text list "Banner_ManIntMsg1": 0 '**Local Message Display**'; 1 '~Spare MB1[0].1'; 2 '~Spare MB1[0].2'; 3 '~Spare MB1[0].3'; 4 '~Spare MB1[0].4'; 5 '~Spare MB1[0].5'; 6 '~Spare MB1[0].6'; 7 '~Spare MB1[0].7'; 8 '~Spare MB1[0].8'; 9 '~Spare MB1[0].9'; 10 '~Spare MB1[0].10'; 11 '~Spare MB1[0].11'; 12 '~Spare MB1[0].12'; 13 '~Spare MB1[0].13'; 14 '~Spare MB1[0].14'; 15 '~Spare MB1[0].15'; 16 '~Spare MB1[0].16'; 17 '~Spare MB1[0].17'; 18 '~Spare MB1[0].18'; 19 '~Spare MB1[0].19'; 20 '~Spare MB1[0].20'; 21 '~Spare MB1[0].21'; 22 '~Spare MB1[0].22'; 23 '~Spare MB1[0].23'; 24 '~Spare MB1[0].24'; 25 '~Spare MB1[0].25'; 26 '~Spare MB1[0].26'; 27 '~Spare MB1[0].27'; 28 '~Spare MB1[0].28'; 29 '~Spare MB1[0].29'; 30 '~Spare MB1[0].30'; 31 '~Spare MB1[0].31'; 32 '~PDPES1 - PDP EtherNet Switch Connection Inhibited MB1[1].0'; 33 '~Spare MB1[1].1'; 34 '~Spare MB1[1].2'; 35 '~MPES1 - Main Panel EtherNet Switch Connection Inhibited MB1[1].3'; 36 '~Spare MB1[1].4'; 37 '~Spare MB1[1].5'; 38 '~MPES2 - Main Panel EtherNet Switch Connection Inhibited MB1[1].6'; 39 '~Spare MB1[1].7'; 40 '~Spare MB1[1].8'; 41 '~MPES3 - Main Panel EtherNet Switch Connection Inhibited MB1[1].9'; 42 '~Spare MB1[1].10'; 43 '~Spare MB1[1].11'; 44 '~S001_004SS1B1 - Service Stand Module Connection Inhibited MB1[1].12'; 45 '~Spare MB1[1].13'; 46 '~Spare MB1[1].14'; 47 '~Spare MB1[1].15'; 48 '~Spare MB1[1].16'; 49 '~MPES1 - Main Panel Control Power Disconnect Not On MB1[1].17'; 50 '~PDP 1 - Panel Output Disconnect Safety Switch Not On MB1[1].18'; 51 '~PDP 2 - Panel Output Disconnect Safety Switch Not On MB1[1].19'; 52 '~PDP 3 - Panel Output Disconnect Safety Switch Not On MB1[1].20'; 53 '~Spare MB1[1].21'; 54 '~Spare MB1[1].22'; 55 '~Spare MB1[1].23'; 56 '~Spare MB1[1].24'; 57 '~Spare MB1[1].25'; 58 '~Spare MB1[1].26'; 59 '~Spare MB1[1].27'; 60 '~Spare MB1[1].28'; 61 '~Spare MB1[1].29'; 62 '~Spare MB1[1].30'; 63 '~Laser Booth-Safe I/O Enclosure Disconnect Safety Switch Not On MB1[1].31'; 64 '~ES1ES1 - ES1 EtherNet Switch Connection Inhibited MB1[2].0'; 65 '~Spare MB1[2].1'; 66 '~Spare MB1[2].2'; 67 '~Spare MB1[2].3'; 68 '~Spare MB1[2].4'; 69 '~Spare MB1[2].5'; 70 '~Spare MB1[2].6'; 71 '~Spare MB1[2].7'; 72 '~Spare MB1[2].8'; 73 '~ES1Sfty - Motion Control Enable Relay #1 MECR1 Still On MB1[2].9'; 74 '~ES1Sfty - Motion Control Enable Relay #1 MECR1 Not On MB1[2].10'; 75 '~ES1Sfty - Motion Control Enable Relay #2 MECR2 Still On MB1[2].11'; 76 '~ES1Sfty - Motion Control Enable Relay #2 MECR2 Not On MB1[2].12'; 77 '~ES1Sfty - EtherNet Switch Sfty Relays RESSR1 RESSR2 Not On MB1[2].13'; 78 '~ES1Sfty - EtherNet Switch Sfty Relays RESSR1 RESSR2 Still On MB1[2].14'; 79 '~Spare MB1[2].15'; 80 '~Spare MB1[2].16'; 81 '~Spare MB1[2].17'; 82 '~Spare MB1[2].18'; 83 '~Spare MB1[2].19'; 84 '~ES1 S001 Safety Gate #1 Open MB1[2].20'; 85 '~ES1 S001 Safety Gate #2 Open MB1[2].21'; 86 '~Spare MB1[2].22'; 87 '~Spare MB1[2].23'; 88 '~Spare MB1[2].24'; 89 '~Spare MB1[2].25'; 90 '~Spare MB1[2].26'; 91 '~Spare MB1[2].27'; 92 '~ES1 S001 Safety Gate #3 Open MB1[2].28'; 93 '~Spare MB1[2].29'; 94 '~Spare MB1[2].30'; 95 '~Spare MB1[2].31'; 96 '~ES2ES1 - ES2 EtherNet Switch Connection Inhibited MB1[3].0'; 97 '~Spare MB1[3].1'; 98 '~Spare MB1[3].2'; 99 '~Spare MB1[3].3'; 100 '~Spare MB1[3].4'; 101 '~Spare MB1[3].5'; 102 '~Spare MB1[3].6'; 103 '~Spare MB1[3].7'; 104 '~Spare MB1[3].8'; 105 '~ES2Sfty - Motion Control Enable Relay #1 MECR1 Still On MB1[3].9'; 106 '~ES2Sfty - Motion Control Enable Relay #1 MECR1 Not On MB1[3].10'; 107 '~ES2Sfty - Motion Control Enable Relay #2 MECR2 Still On MB1[3].11'; 108 '~ES2Sfty - Motion Control Enable Relay #2 MECR2 Not On MB1[3].12'; 109 '~ES2Sfty - EtherNet Switch Sfty Relays RESSR1 RESSR2 Not On MB1[3].13'; 110 '~ES2Sfty - EtherNet Switch Sfty Relays RESSR1 RESSR2 Still On MB1[3].14'; 111 '~Spare MB1[3].15'; 112 '~Spare MB1[3].16'; 113 '~Spare MB1[3].17'; 114 '~Spare MB1[3].18'; 115 '~Spare MB1[3].19'; 116 '~ES2 S001 Safety Gate #1 Open MB1[3].20'; 117 '~ES2 S001 Safety Gate #2 Open MB1[3].21'; 118 '~Spare MB1[3].22'; 119 '~Spare MB1[3].23'; 120 '~Spare MB1[3].24'; 121 '~Spare MB1[3].25'; 122 '~Spare MB1[3].26'; 123 '~Spare MB1[3].27'; 124 '~Spare MB1[3].28'; 125 '~Spare MB1[3].29'; 126 '~Spare MB1[3].30'; 127 '~Spare MB1[3].31'; 128 '~PV1ES1 - PV1 EtherNet Switch Connection Inhibited MB1[4].0'; 129 '~Spare MB1[4].1'; 130 '~Spare MB1[4].2'; 131 '~Spare MB1[4].3'; 132 '~Spare MB1[4].4'; 133 '~Spare MB1[4].5'; 134 '~Spare MB1[4].6'; 135 '~Spare MB1[4].7'; 136 '~Spare MB1[4].8'; 137 '~Spare MB1[4].9'; 138 '~Spare MB1[4].10'; 139 '~PV1Sfty - EtherNet Switch Sfty Relays RESSR1 RESSR2 Not On MB1[4].11'; 140 '~PV1Sfty - EtherNet Switch Sfty Relays RESSR1 RESSR2 Still On MB1[4].12'; 141 '~Spare MB1[4].13'; 142 '~Spare MB1[4].14'; 143 '~PV1 S001 E-Stop Depressed MB1[4].15'; 144 '~PV1 S001 Safety Gate #1 Open MB1[4].16'; 145 '~PV1 S001 Safety Gate #2 Open MB1[4].17'; 146 '~PV1 S001 Safety Gate #3 Open MB1[4].18'; 147 '~Spare MB1[4].19'; 148 '~Spare MB1[4].20'; 149 '~Spare MB1[4].21'; 150 '~Spare MB1[4].22'; 151 '~Spare MB1[4].23'; 152 '~S001 Both PanelViews Have Manual Selected MB1[4].24'; 153 '~S001 PanelView 1 Manual Selected MB1[4].25'; 154 '~Spare MB1[4].26'; 155 '~Spare MB1[4].27'; 156 '~PV1 S001 Auto Not Selected MB1[4].28'; 157 '~PV1 S001 Not In Auto Or Manual MB1[4].29'; 158 '~Spare MB1[4].30'; 159 '~Spare MB1[4].31'; 160 '~PV2ES1 - PV2 EtherNet Switch Connection Inhibited MB1[5].0'; 161 '~Spare MB1[5].1'; 162 '~Spare MB1[5].2'; 163 '~Spare MB1[5].3'; 164 '~Spare MB1[5].4'; 165 '~Spare MB1[5].5'; 166 '~Spare MB1[5].6'; 167 '~Spare MB1[5].7'; 168 '~Spare MB1[5].8'; 169 '~Spare MB1[5].9'; 170 '~Spare MB1[5].10'; 171 '~PV2Sfty - EtherNet Switch Sfty Relays RESSR1 RESSR2 Not On MB1[5].11'; 172 '~PV2Sfty - EtherNet Switch Sfty Relays RESSR1 RESSR2 Still On MB1[5].12'; 173 '~Spare MB1[5].13'; 174 '~Spare MB1[5].14'; 175 '~PV2 S001 E-Stop Depressed MB1[5].15'; 176 '~PV2 S001 Safety Gate #1 Open MB1[5].16'; 177 '~PV2 S001 Safety Gate #2 Open MB1[5].17'; 178 '~PV2 S001 Safety Gate #3 Open MB1[5].18'; 179 '~Spare MB1[5].19'; 180 '~Spare MB1[5].20'; 181 '~Spare MB1[5].21'; 182 '~Spare MB1[5].22'; 183 '~Spare MB1[5].23'; 184 '~Spare MB1[5].24'; 185 '~S001 PanelView 2 Manual Selected MB1[5].25'; 186 '~Spare MB1[5].26'; 187 '~Spare MB1[5].27'; 188 '~PV2 S001 Auto Not Selected MB1[5].28'; 189 '~PV2 S001 Not In Auto Or Manual MB1[5].29'; 190 '~Spare MB1[5].30'; 191 '~Spare MB1[5].31'; 192 '~S001R01ES1 - S001R01 EtherNet Switch Connection Inhibited MB1[6].0'; 193 '~Spare MB1[6].1'; 194 '~Spare MB1[6].2'; 195 '~Spare MB1[6].3'; 196 '~Spare MB1[6].4'; 197 '~Spare MB1[6].5'; 198 '~Spare MB1[6].6'; 199 '~Spare MB1[6].7'; 200 '~Spare MB1[6].8'; 201 '~Spare MB1[6].9'; 202 '~Spare MB1[6].10'; 203 '~Spare MB1[6].11'; 204 '~Spare MB1[6].12'; 205 '~Spare MB1[6].13'; 206 '~Spare MB1[6].14'; 207 '~Spare MB1[6].15'; 208 '~Spare MB1[6].16'; 209 '~S001R01Sfty - Robot E-Stop Depressed MB1[6].17'; 210 '~S001R01Sfty - Robot Safety Interface Not Enabled MB1[6].18'; 211 '~S001R01Sfty - Robot DCS Has Been Edited MB1[6].19'; 212 '~S001R01CN - Robot Controller Connection Inhibited MB1[6].20'; 213 '~S001R01E#B# - Robot End Effector Module Connection Inhibited MB1[6].21'; 214 '~S001R01E#B# - Robot End Effector Module Connection Inhibited MB1[6].22'; 215 '~S001R01E#B# - Robot End Effector Module Connection Inhibited MB1[6].23'; 216 '~S001R01E#B# - Robot End Effector Module Connection Inhibited MB1[6].24'; 217 '~S001R01E#B# - Robot End Effector Module Connection Inhibited MB1[6].25'; 218 '~S001R01E#B# - Robot End Effector Module Connection Inhibited MB1[6].26'; 219 '~S001R01E#B# - Robot End Effector Module Connection Inhibited MB1[6].27'; 220 '~S001R01E#B# - Robot End Effector Module Connection Inhibited MB1[6].28'; 221 '~S001R01E#B# - Robot End Effector Module Connection Inhibited MB1[6].29'; 222 '~Spare MB1[6].30'; 223 '~Spare MB1[6].31'; 224 '~Spare MB1[7].0'; 225 '~S001R01F#B# - Robot Process I/O Connection Inhibited MB1[7].1'; 226 '~S001R01F#B# - Robot Process I/O Connection Inhibited MB1[7].2'; 227 '~S001R01F#B# - Robot Process I/O Connection Inhibited MB1[7].3'; 228 '~S001R01F#B# - Robot Process I/O Connection Inhibited MB1[7].4'; 229 '~Spare MB1[7].5'; 230 '~Spare MB1[7].6'; 231 '~Spare MB1[7].7'; 232 '~Spare MB1[7].8'; 233 '~Spare MB1[7].9'; 234 '~S001R01CN.I.Safety - Chain Fault MB1[7].10'; 235 '~S001R01CN.I.AirOn - Robot Air Not On MB1[7].11'; 236 '~S001R01CN.I.RbtAuto - Robot Not in Auto MB1[7].12'; 237 '~S001R01CN.M.InTeach - Robot In Teach MB1[7].13'; 238 '~S001R01CN.I.AtMaintPos - Robot At Maintenace MB1[7].14'; 239 '~S001R01CN.I.RunEnblInterruptAck - Robot In Hold MB1[7].15'; 240 '~S001R01CN.M.MaintPosSeld - Robot Maintenance Selected MB1[7].16'; 241 '~Spare MB1[7].17'; 242 '~Spare MB1[7].18'; 243 '~Spare MB1[7].19'; 244 '~S001R01CN.I.ExtAppCommFlt - Robot Application Communication Fault MB1[7].20'; 245 '~S001R01CN.M.AbortPickupSeld - Robot Abort Pickup Selected MB1[7].21'; 246 '~S001R01CN.M.RetFmPounceSeld - Robot Return From Pounce Selected MB1[7].22'; 247 '~S001R01CN.I.StudWld1 Comm Not OK MB1[7].23'; 248 '~S001R01CN.I.StudWld2 Comm Not OK MB1[7].24'; 249 '~S001R01CN.I.WldMode - Robot In No Weld MB1[7].25'; 250 '~S001R01CN.I.PulledTipBypSS - Robot Pulled Tip Bypass Selected MB1[7].26'; 251 '~S001R01CN.I.FlowNoFlowSS - Robot In No Flow MB1[7].27'; 252 '~S001R01CN.I.RvtNoRvtSS - Robot In No Rivet MB1[7].28'; 253 '~S001R01CN.I.WldCtrlCommOk1 - Robot Weld Controller 1 Comm Not OK MB1[7].29'; 254 '~S001R01CN.I.WldModeStud - Robot In No Weld Stud MB1[7].30'; 255 '~S001R01CN.Ix.MigWldNoWld - Robot In No Weld Mig MB1[7].31'; 256 '~S001R01CN.I.StudWld1Rdy - Robot Stud Weld Controller 1 Not Ready MB1[8].0'; 257 '~S001R01CN.I.Rvt1RdyToOperate - Robot Rivet Controller 1 Not Ready MB1[8].1'; 258 '~S001R01CN.Ix.MigRdy - Robot Mig Weld Controller Not Ready MB1[8].2'; 259 '~S001R01CN.Ix.MigWldNoWld - Robot In No Weld MB1[8].3'; 260 '~Spare MB1[8].4'; 261 '~S001R01CN.I.WldCtrlCommOk2 - Robot Weld Controller 2 Comm Not OK MB1[8].5'; 262 '~Spare MB1[8].6'; 263 '~Spare MB1[8].7'; 264 '~S001R01CN.I.StudWld2Rdy - Robot Stud Weld Controller 2 Not Ready MB1[8].8'; 265 '~S001R01CN.I.Rvt2RdyToOperate - Robot Rivet Controller 2 Not Ready MB1[8].9'; 266 '~S001R01CN.Ix.LaserWldOn - Robot Laser In No Cut MB1[8].10'; 267 '~S001R01CN.Ix.GlassNotPres - Robot Laser Glass Not Present MB1[8].11'; 268 '~S001R01CN.Ix.LaserHeadRdy - Robot Laser Head Not Ready MB1[8].12'; 269 '~S001R01CN.Ix.ChillerOn - Robot Laser Chiller Not On MB1[8].13'; 270 '~S001R01CN.Ix.GasOn - Robot Gas Not On MB1[8].14'; 271 '~S001R01 Power Meter Not Ready MB1[8].15'; 272 '~S001R01 No Wire Present Replace Barrel MB1[8].16'; 273 '~S001R01 Wire Feeder Fault Timer MB1[8].17'; 274 '~S001R01CN.Ix.NRFlt - Robot Nut Runner Not Ready MB1[8].18'; 275 '~Spare MB1[8].19'; 276 '~S001R01CN.M.WrongRivetAtNose - Remove Wrong Rivet At Nose MB1[8].20'; 277 '~S001R01CN.M.DisableRbtDrvs - In Rivet Zone But Riveter Not In Auto MB1[8].21'; 278 '~S001R01CN.I.Rvt1SystemInAuto - Rivet Controller 1 Not In Auto MB1[8].22'; 279 '~S001R01CN.I.Rvt2SystemInAuto - Rivet Controller 2 Not In Auto MB1[8].23'; 280 '~S001R01CN.M.RvtC1ReelCtr.DN - Reel Change Required MB1[8].24'; 281 '~S001R01CN.M.RvtC2ReelCtr.DN - Reel Change Required MB1[8].25'; 282 '~S001R01CN.M.AbortSkipRemain - SkipRemaining Aborted, Reset At Rbt Controller Is Required MB1[8].26'; 283 '~Spare MB1[8].27'; 284 '~Spare MB1[8].28'; 285 '~Spare MB1[8].29'; 286 '~Spare MB1[8].30'; 287 '~Spare MB1[8].31'; 288 '~Spare MB1[9].0'; 289 '~Spare MB1[9].1'; 290 '~Spare MB1[9].2'; 291 '~Spare MB1[9].3'; 292 '~Spare MB1[9].4'; 293 '~Spare MB1[9].5'; 294 '~Spare MB1[9].6'; 295 '~Spare MB1[9].7'; 296 '~Spare MB1[9].8'; 297 '~Spare MB1[9].9'; 298 '~Spare MB1[9].10'; 299 '~Spare MB1[9].11'; 300 '~Spare MB1[9].12'; 301 '~Spare MB1[9].13'; 302 '~Spare MB1[9].14'; 303 '~Spare MB1[9].15'; 304 '~Spare MB1[9].16'; 305 '~Spare MB1[9].17'; 306 '~Spare MB1[9].18'; 307 '~Spare MB1[9].19'; 308 '~Spare MB1[9].20'; 309 '~Spare MB1[9].21'; 310 '~Spare MB1[9].22'; 311 '~Spare MB1[9].23'; 312 '~Spare MB1[9].24'; 313 '~Spare MB1[9].25'; 314 '~Spare MB1[9].26'; 315 '~Spare MB1[9].27'; 316 '~Spare MB1[9].28'; 317 '~Spare MB1[9].29'; 318 '~Spare MB1[9].30'; 319 '~Spare MB1[9].31'; 320 '~Spare MB1[10].0'; 321 '~Spare MB1[10].1'; 322 '~Spare MB1[10].2'; 323 '~Spare MB1[10].3'; 324 '~Spare MB1[10].4'; 325 '~Spare MB1[10].5'; 326 '~Spare MB1[10].6'; 327 '~Spare MB1[10].7'; 328 '~Spare MB1[10].8'; 329 '~Spare MB1[10].9'; 330 '~Spare MB1[10].10'; 331 '~Spare MB1[10].11'; 332 '~Spare MB1[10].12'; 333 '~Spare MB1[10].13'; 334 '~Spare MB1[10].14'; 335 '~Spare MB1[10].15'; 336 '~Spare MB1[10].16'; 337 '~Spare MB1[10].17'; 338 '~Spare MB1[10].18'; 339 '~Spare MB1[10].19'; 340 '~Spare MB1[10].20'; 341 '~Spare MB1[10].21'; 342 '~Spare MB1[10].22'; 343 '~Spare MB1[10].23'; 344 '~Spare MB1[10].24'; 345 '~Spare MB1[10].25'; 346 '~Spare MB1[10].26'; 347 '~Spare MB1[10].27'; 348 '~Spare MB1[10].28'; 349 '~Spare MB1[10].29'; 350 '~Spare MB1[10].30'; 351 '~Spare MB1[10].31'; 352 '~Spare MB1[11].0'; 353 '~Spare MB1[11].1'; 354 '~Spare MB1[11].2'; 355 '~Spare MB1[11].3'; 356 '~Spare MB1[11].4'; 357 '~Spare MB1[11].5'; 358 '~Spare MB1[11].6'; 359 '~Spare MB1[11].7'; 360 '~Spare MB1[11].8'; 361 '~Spare MB1[11].9'; 362 '~Spare MB1[11].10'; 363 '~Spare MB1[11].11'; 364 '~Spare MB1[11].12'; 365 '~Spare MB1[11].13'; 366 '~Spare MB1[11].14'; 367 '~Spare MB1[11].15'; 368 '~Spare MB1[11].16'; 369 '~Spare MB1[11].17'; 370 '~Spare MB1[11].18'; 371 '~Spare MB1[11].19'; 372 '~Spare MB1[11].20'; 373 '~Spare MB1[11].21'; 374 '~Spare MB1[11].22'; 375 '~Spare MB1[11].23'; 376 '~Spare MB1[11].24'; 377 '~Spare MB1[11].25'; 378 '~Spare MB1[11].26'; 379 '~Spare MB1[11].27'; 380 '~Spare MB1[11].28'; 381 '~Spare MB1[11].29'; 382 '~Spare MB1[11].30'; 383 '~Spare MB1[11].31'; 384 '~S001R02ES1 - S001R02 EtherNet Switch Connection Inhibited MB1[12].0'; 385 '~Spare MB1[12].1'; 386 '~Spare MB1[12].2'; 387 '~Spare MB1[12].3'; 388 '~Spare MB1[12].4'; 389 '~Spare MB1[12].5'; 390 '~Spare MB1[12].6'; 391 '~Spare MB1[12].7'; 392 '~Spare MB1[12].8'; 393 '~Spare MB1[12].9'; 394 '~Spare MB1[12].10'; 395 '~Spare MB1[12].11'; 396 '~Spare MB1[12].12'; 397 '~Spare MB1[12].13'; 398 '~Spare MB1[12].14'; 399 '~Spare MB1[12].15'; 400 '~Spare MB1[12].16'; 401 '~S001R02Sfty - Robot E-Stop Depressed MB1[12].17'; 402 '~S001R02Sfty - Robot Safety Interface Not Enabled MB1[12].18'; 403 '~S001R02Sfty - Robot DCS Has Been Edited MB1[12].19'; 404 '~S001R02CN - Robot Controller Connection Inhibited MB1[12].20'; 405 '~S001R02E#B# - Robot End Effector Module Connection Inhibited MB1[12].21'; 406 '~S001R02E#B# - Robot End Effector Module Connection Inhibited MB1[12].22'; 407 '~S001R02E#B# - Robot End Effector Module Connection Inhibited MB1[12].23'; 408 '~S001R02E#B# - Robot End Effector Module Connection Inhibited MB1[12].24'; 409 '~S001R02E#B# - Robot End Effector Module Connection Inhibited MB1[12].25'; 410 '~S001R02E#B# - Robot End Effector Module Connection Inhibited MB1[12].26'; 411 '~S001R02E#B# - Robot End Effector Module Connection Inhibited MB1[12].27'; 412 '~S001R02E#B# - Robot End Effector Module Connection Inhibited MB1[12].28'; 413 '~S001R02E#B# - Robot End Effector Module Connection Inhibited MB1[12].29'; 414 '~Spare MB1[12].30'; 415 '~Spare MB1[12].31'; 416 '~Spare MB1[13].0'; 417 '~S001R02F#B# - Robot Process I/O Connection Inhibited MB1[13].1'; 418 '~S001R02F#B# - Robot Process I/O Connection Inhibited MB1[13].2'; 419 '~S001R02F#B# - Robot Process I/O Connection Inhibited MB1[13].3'; 420 '~S001R02F#B# - Robot Process I/O Connection Inhibited MB1[13].4'; 421 '~Spare MB1[13].5'; 422 '~Spare MB1[13].6'; 423 '~Spare MB1[13].7'; 424 '~Spare MB1[13].8'; 425 '~Spare MB1[13].9'; 426 '~S001R02CN.I.Safety - Chain Fault MB1[13].10'; 427 '~S001R02CN.I.AirOn - Robot Air Not On MB1[13].11'; 428 '~S001R02CN.I.RbtAuto - Robot Not in Auto MB1[13].12'; 429 '~S001R02CN.M.InTeach - Robot In Teach MB1[13].13'; 430 '~S001R02CN.I.AtMaintPos - Robot At Maintenace MB1[13].14'; 431 '~S001R02CN.I.RunEnblInterruptAck - Robot In Hold MB1[13].15'; 432 '~S001R02CN.M.MaintPosSeld - Robot Maintenance Selected MB1[13].16'; 433 '~Spare MB1[13].17'; 434 '~Spare MB1[13].18'; 435 '~Spare MB1[13].19'; 436 '~S001R02CN.I.ExtAppCommFlt - Robot Application Communication Fault MB1[13].20'; 437 '~S001R02CN.M.AbortPickupSeld - Robot Abort Pickup Selected MB1[13].21'; 438 '~S001R02CN.M.RetFmPounceSeld - Robot Return From Pounce Selected MB1[13].22'; 439 '~S001R02CN.I.StudWld1 Comm Not OK MB1[13].23'; 440 '~S001R02CN.I.StudWld2 Comm Not OK MB1[13].24'; 441 '~S001R02CN.I.WldMode - Robot In No Weld MB1[13].25'; 442 '~S001R02CN.I.PulledTipBypSS - Robot Pulled Tip Bypass Selected MB1[13].26'; 443 '~S001R02CN.I.FlowNoFlowSS - Robot In No Flow MB1[13].27'; 444 '~S001R02CN.I.RvtNoRvtSS - Robot In No Rivet MB1[13].28'; 445 '~S001R02CN.I.WldCtrlCommOk1 - Robot Weld Controller 1 Comm Not OK MB1[13].29'; 446 '~S001R02CN.I.WldModeStud - Robot In No Weld Stud MB1[13].30'; 447 '~S001R02CN.Ix.MigWldNoWld - Robot In No Weld Mig MB1[13].31'; 448 '~S001R02CN.I.StudWld1Rdy - Robot Stud Weld Controller 1 Not Ready MB1[14].0'; 449 '~S001R02CN.I.Rvt1RdyToOperate - Robot Rivet Controller 1 Not Ready MB1[14].1'; 450 '~S001R02CN.Ix.MigRdy - Robot Mig Weld Controller Not Ready MB1[14].2'; 451 '~S001R02CN.Ix.MigWldNoWld - Robot In No Weld MB1[14].3'; 452 '~Spare MB1[14].4'; 453 '~S001R02CN.I.WldCtrlCommOk2 - Robot Weld Controller 2 Comm Not OK MB1[14].5'; 454 '~Spare MB1[14].6'; 455 '~Spare MB1[14].7'; 456 '~S001R02CN.I.StudWld2Rdy - Robot Stud Weld Controller 2 Not Ready MB1[14].8'; 457 '~S001R02CN.I.Rvt2RdyToOperate - Robot Rivet Controller 2 Not Ready MB1[14].9'; 458 '~S001R02CN.Ix.LaserWldOn - Robot Laser In No Cut MB1[14].10'; 459 '~S001R02CN.Ix.GlassNotPres - Robot Laser Glass Not Present MB1[14].11'; 460 '~S001R02CN.Ix.LaserHeadRdy - Robot Laser Head Not Ready MB1[14].12'; 461 '~S001R02CN.Ix.ChillerOn - Robot Laser Chiller Not On MB1[14].13'; 462 '~S001R02CN.Ix.GasOn - Robot Gas Not On MB1[14].14'; 463 '~S001R02 Power Meter Not Ready MB1[14].15'; 464 '~S001R02 No Wire Present Replace Barrel MB1[14].16'; 465 '~S001R02 Wire Feeder Fault Timer MB1[14].17'; 466 '~S001R02CN.Ix.NRFlt - Robot Nut Runner Not Ready MB1[14].18'; 467 '~Spare MB1[14].19'; 468 '~S001R02CN.M.WrongRivetAtNose - Remove Wrong Rivet At Nose MB1[14].20'; 469 '~S001R02CN.M.DisableRbtDrvs - In Rivet Zone But Riveter Not In Auto MB1[14].21'; 470 '~S001R02CN.I.Rvt1SystemInAuto - Rivet Controller 1 Not In Auto MB1[14].22'; 471 '~S001R02CN.I.Rvt2SystemInAuto - Rivet Controller 2 Not In Auto MB1[14].23'; 472 '~S001R02CN.M.RvtC1ReelCtr.DN - Reel Change Required MB1[14].24'; 473 '~S001R02CN.M.RvtC2ReelCtr.DN - Reel Change Required MB1[14].25'; 474 '~S001R02CN.M.AbortSkipRemain - SkipRemaining Aborted, Reset At Rbt Controller Is Required MB1[14].26'; 475 '~Spare MB1[14].27'; 476 '~Spare MB1[14].28'; 477 '~Spare MB1[14].29'; 478 '~Spare MB1[14].30'; 479 '~Spare MB1[14].31'; 480 '~Spare MB1[15].0'; 481 '~Spare MB1[15].1'; 482 '~Spare MB1[15].2'; 483 '~Spare MB1[15].3'; 484 '~Spare MB1[15].4'; 485 '~Spare MB1[15].5'; 486 '~Spare MB1[15].6'; 487 '~Spare MB1[15].7'; 488 '~Spare MB1[15].8'; 489 '~Spare MB1[15].9'; 490 '~Spare MB1[15].10'; 491 '~Spare MB1[15].11'; 492 '~Spare MB1[15].12'; 493 '~Spare MB1[15].13'; 494 '~Spare MB1[15].14'; 495 '~Spare MB1[15].15'; 496 '~Spare MB1[15].16'; 497 '~Spare MB1[15].17'; 498 '~Spare MB1[15].18'; 499 '~Spare MB1[15].19'; 500 '~Spare MB1[15].20'; 501 '~Spare MB1[15].21'; 502 '~Spare MB1[15].22'; 503 '~Spare MB1[15].23'; 504 '~Spare MB1[15].24'; 505 '~Spare MB1[15].25'; 506 '~Spare MB1[15].26'; 507 '~Spare MB1[15].27'; 508 '~Spare MB1[15].28'; 509 '~Spare MB1[15].29'; 510 '~Spare MB1[15].30'; 511 '~Spare MB1[15].31'; 512 '~Spare MB1[16].0'; 513 '~Spare MB1[16].1'; 514 '~Spare MB1[16].2'; 515 '~Spare MB1[16].3'; 516 '~Spare MB1[16].4'; 517 '~Spare MB1[16].5'; 518 '~Spare MB1[16].6'; 519 '~Spare MB1[16].7'; 520 '~Spare MB1[16].8'; 521 '~Spare MB1[16].9'; 522 '~Spare MB1[16].10'; 523 '~Spare MB1[16].11'; 524 '~Spare MB1[16].12'; 525 '~Spare MB1[16].13'; 526 '~Spare MB1[16].14'; 527 '~Spare MB1[16].15'; 528 '~Spare MB1[16].16'; 529 '~Spare MB1[16].17'; 530 '~Spare MB1[16].18'; 531 '~Spare MB1[16].19'; 532 '~Spare MB1[16].20'; 533 '~Spare MB1[16].21'; 534 '~Spare MB1[16].22'; 535 '~Spare MB1[16].23'; 536 '~Spare MB1[16].24'; 537 '~Spare MB1[16].25'; 538 '~Spare MB1[16].26'; 539 '~Spare MB1[16].27'; 540 '~Spare MB1[16].28'; 541 '~Spare MB1[16].29'; 542 '~Spare MB1[16].30'; 543 '~Spare MB1[16].31'; 544 '~Spare MB1[17].0'; 545 '~Spare MB1[17].1'; 546 '~Spare MB1[17].2'; 547 '~Spare MB1[17].3'; 548 '~Spare MB1[17].4'; 549 '~Spare MB1[17].5'; 550 '~Spare MB1[17].6'; 551 '~Spare MB1[17].7'; 552 '~Spare MB1[17].8'; 553 '~Spare MB1[17].9'; 554 '~Spare MB1[17].10'; 555 '~Spare MB1[17].11'; 556 '~Spare MB1[17].12'; 557 '~Spare MB1[17].13'; 558 '~Spare MB1[17].14'; 559 '~Spare MB1[17].15'; 560 '~Spare MB1[17].16'; 561 '~Spare MB1[17].17'; 562 '~Spare MB1[17].18'; 563 '~Spare MB1[17].19'; 564 '~Spare MB1[17].20'; 565 '~Spare MB1[17].21'; 566 '~Spare MB1[17].22'; 567 '~Spare MB1[17].23'; 568 '~Spare MB1[17].24'; 569 '~Spare MB1[17].25'; 570 '~Spare MB1[17].26'; 571 '~Spare MB1[17].27'; 572 '~Spare MB1[17].28'; 573 '~Spare MB1[17].29'; 574 '~Spare MB1[17].30'; 575 '~Spare MB1[17].31'; 576 '~S001R03ES1 - S001R03 EtherNet Switch Connection Inhibited MB1[18].0'; 577 '~Spare MB1[18].1'; 578 '~Spare MB1[18].2'; 579 '~Spare MB1[18].3'; 580 '~Spare MB1[18].4'; 581 '~Spare MB1[18].5'; 582 '~Spare MB1[18].6'; 583 '~Spare MB1[18].7'; 584 '~Spare MB1[18].8'; 585 '~Spare MB1[18].9'; 586 '~Spare MB1[18].10'; 587 '~Spare MB1[18].11'; 588 '~Spare MB1[18].12'; 589 '~Spare MB1[18].13'; 590 '~Spare MB1[18].14'; 591 '~Spare MB1[18].15'; 592 '~Spare MB1[18].16'; 593 '~S001R03Sfty - Robot E-Stop Depressed MB1[18].17'; 594 '~S001R03Sfty - Robot Safety Interface Not Enabled MB1[18].18'; 595 '~S001R03Sfty - Robot DCS Has Been Edited MB1[18].19'; 596 '~S001R03CN - Robot Controller Connection Inhibited MB1[18].20'; 597 '~S001R03E#B# - Robot End Effector Module Connection Inhibited MB1[18].21'; 598 '~S001R03E#B# - Robot End Effector Module Connection Inhibited MB1[18].22'; 599 '~S001R03E#B# - Robot End Effector Module Connection Inhibited MB1[18].23'; 600 '~S001R03E#B# - Robot End Effector Module Connection Inhibited MB1[18].24'; 601 '~S001R03E#B# - Robot End Effector Module Connection Inhibited MB1[18].25'; 602 '~S001R03E#B# - Robot End Effector Module Connection Inhibited MB1[18].26'; 603 '~S001R03E#B# - Robot End Effector Module Connection Inhibited MB1[18].27'; 604 '~S001R03E#B# - Robot End Effector Module Connection Inhibited MB1[18].28'; 605 '~S001R03E#B# - Robot End Effector Module Connection Inhibited MB1[18].29'; 606 '~Spare MB1[18].30'; 607 '~Spare MB1[18].31'; 608 '~Spare MB1[19].0'; 609 '~S001R03F#B# - Robot Process I/O Connection Inhibited MB1[19].1'; 610 '~S001R03F#B# - Robot Process I/O Connection Inhibited MB1[19].2'; 611 '~S001R03F#B# - Robot Process I/O Connection Inhibited MB1[19].3'; 612 '~S001R03F#B# - Robot Process I/O Connection Inhibited MB1[19].4'; 613 '~Spare MB1[19].5'; 614 '~Spare MB1[19].6'; 615 '~Spare MB1[19].7'; 616 '~Spare MB1[19].8'; 617 '~Spare MB1[19].9'; 618 '~S001R03CN.I.Safety - Chain Fault MB1[19].10'; 619 '~S001R03CN.I.AirOn - Robot Air Not On MB1[19].11'; 620 '~S001R03CN.I.RbtAuto - Robot Not in Auto MB1[19].12'; 621 '~S001R03CN.M.InTeach - Robot In Teach MB1[19].13'; 622 '~S001R03CN.I.AtMaintPos - Robot At Maintenace MB1[19].14'; 623 '~S001R03CN.I.RunEnblInterruptAck - Robot In Hold MB1[19].15'; 624 '~S001R03CN.M.MaintPosSeld - Robot Maintenance Selected MB1[19].16'; 625 '~Spare MB1[19].17'; 626 '~Spare MB1[19].18'; 627 '~Spare MB1[19].19'; 628 '~S001R03CN.I.ExtAppCommFlt - Robot Application Communication Fault MB1[19].20'; 629 '~S001R03CN.M.AbortPickupSeld - Robot Abort Pickup Selected MB1[19].21'; 630 '~S001R03CN.M.RetFmPounceSeld - Robot Return From Pounce Selected MB1[19].22'; 631 '~S001R03CN.I.StudWld1 Comm Not OK MB1[19].23'; 632 '~S001R03CN.I.StudWld2 Comm Not OK MB1[19].24'; 633 '~S001R03CN.I.WldMode - Robot In No Weld MB1[19].25'; 634 '~S001R03CN.I.PulledTipBypSS - Robot Pulled Tip Bypass Selected MB1[19].26'; 635 '~S001R03CN.I.FlowNoFlowSS - Robot In No Flow MB1[19].27'; 636 '~S001R03CN.I.RvtNoRvtSS - Robot In No Rivet MB1[19].28'; 637 '~S001R03CN.I.WldCtrlCommOk1 - Robot Weld Controller 1 Comm Not OK MB1[19].29'; 638 '~S001R03CN.I.WldModeStud - Robot In No Weld Stud MB1[19].30'; 639 '~S001R03CN.Ix.MigWldNoWld - Robot In No Weld Mig MB1[19].31'; 640 '~S001R03CN.I.StudWld1Rdy - Robot Stud Weld Controller 1 Not Ready MB1[20].0'; 641 '~S001R03CN.I.Rvt1RdyToOperate - Robot Rivet Controller 1 Not Ready MB1[20].1'; 642 '~S001R03CN.Ix.MigRdy - Robot Mig Weld Controller Not Ready MB1[20].2'; 643 '~S001R03CN.Ix.MigWldNoWld - Robot In No Weld MB1[20].3'; 644 '~Spare MB1[20].4'; 645 '~S001R03CN.I.WldCtrlCommOk2 - Robot Weld Controller 2 Comm Not OK MB1[20].5'; 646 '~Spare MB1[20].6'; 647 '~Spare MB1[20].7'; 648 '~S001R03CN.I.StudWld2Rdy - Robot Stud Weld Controller 2 Not Ready MB1[20].8'; 649 '~S001R03CN.I.Rvt2RdyToOperate - Robot Rivet Controller 2 Not Ready MB1[20].9'; 650 '~S001R03CN.Ix.LaserWldOn - Robot Laser In No Cut MB1[20].10'; 651 '~S001R03CN.Ix.GlassNotPres - Robot Laser Glass Not Present MB1[20].11'; 652 '~S001R03CN.Ix.LaserHeadRdy - Robot Laser Head Not Ready MB1[20].12'; 653 '~S001R03CN.Ix.ChillerOn - Robot Laser Chiller Not On MB1[20].13'; 654 '~S001R03CN.Ix.GasOn - Robot Gas Not On MB1[20].14'; 655 '~S001R03 Power Meter Not Ready MB1[20].15'; 656 '~S001R03 No Wire Present Replace Barrel MB1[20].16'; 657 '~S001R03 Wire Feeder Fault Timer MB1[20].17'; 658 '~S001R03CN.Ix.NRFlt - Robot Nut Runner Not Ready MB1[20].18'; 659 '~Spare MB1[20].19'; 660 '~S001R03CN.M.WrongRivetAtNose - Remove Wrong Rivet At Nose MB1[20].20'; 661 '~S001R03CN.M.DisableRbtDrvs - In Rivet Zone But Riveter Not In Auto MB1[20].21'; 662 '~S001R03CN.I.Rvt1SystemInAuto - Rivet Controller 1 Not In Auto MB1[20].22'; 663 '~S001R03CN.I.Rvt2SystemInAuto - Rivet Controller 2 Not In Auto MB1[20].23'; 664 '~S001R03CN.M.RvtC1ReelCtr.DN - Reel Change Required MB1[20].24'; 665 '~S001R03CN.M.RvtC2ReelCtr.DN - Reel Change Required MB1[20].25'; 666 '~S001R03CN.M.AbortSkipRemain - SkipRemaining Aborted, Reset At Rbt Controller Is Required MB1[20].26'; 667 '~Spare MB1[20].27'; 668 '~Spare MB1[20].28'; 669 '~Spare MB1[20].29'; 670 '~Spare MB1[20].30'; 671 '~Spare MB1[20].31'; 672 '~Spare MB1[21].0'; 673 '~Spare MB1[21].1'; 674 '~Spare MB1[21].2'; 675 '~Spare MB1[21].3'; 676 '~Spare MB1[21].4'; 677 '~Spare MB1[21].5'; 678 '~Spare MB1[21].6'; 679 '~Spare MB1[21].7'; 680 '~Spare MB1[21].8'; 681 '~Spare MB1[21].9'; 682 '~Spare MB1[21].10'; 683 '~Spare MB1[21].11'; 684 '~Spare MB1[21].12'; 685 '~Spare MB1[21].13'; 686 '~Spare MB1[21].14'; 687 '~Spare MB1[21].15'; 688 '~Spare MB1[21].16'; 689 '~Spare MB1[21].17'; 690 '~Spare MB1[21].18'; 691 '~Spare MB1[21].19'; 692 '~Spare MB1[21].20'; 693 '~Spare MB1[21].21'; 694 '~Spare MB1[21].22'; 695 '~Spare MB1[21].23'; 696 '~Spare MB1[21].24'; 697 '~Spare MB1[21].25'; 698 '~Spare MB1[21].26'; 699 '~Spare MB1[21].27'; 700 '~Spare MB1[21].28'; 701 '~Spare MB1[21].29'; 702 '~Spare MB1[21].30'; 703 '~Spare MB1[21].31'; 704 '~Spare MB1[22].0'; 705 '~Spare MB1[22].1'; 706 '~Spare MB1[22].2'; 707 '~Spare MB1[22].3'; 708 '~Spare MB1[22].4'; 709 '~Spare MB1[22].5'; 710 '~Spare MB1[22].6'; 711 '~Spare MB1[22].7'; 712 '~Spare MB1[22].8'; 713 '~Spare MB1[22].9'; 714 '~Spare MB1[22].10'; 715 '~Spare MB1[22].11'; 716 '~Spare MB1[22].12'; 717 '~Spare MB1[22].13'; 718 '~Spare MB1[22].14'; 719 '~Spare MB1[22].15'; 720 '~Spare MB1[22].16'; 721 '~Spare MB1[22].17'; 722 '~Spare MB1[22].18'; 723 '~Spare MB1[22].19'; 724 '~Spare MB1[22].20'; 725 '~Spare MB1[22].21'; 726 '~Spare MB1[22].22'; 727 '~Spare MB1[22].23'; 728 '~Spare MB1[22].24'; 729 '~Spare MB1[22].25'; 730 '~Spare MB1[22].26'; 731 '~Spare MB1[22].27'; 732 '~Spare MB1[22].28'; 733 '~Spare MB1[22].29'; 734 '~Spare MB1[22].30'; 735 '~Spare MB1[22].31'; 736 '~Spare MB1[23].0'; 737 '~Spare MB1[23].1'; 738 '~Spare MB1[23].2'; 739 '~Spare MB1[23].3'; 740 '~Spare MB1[23].4'; 741 '~Spare MB1[23].5'; 742 '~Spare MB1[23].6'; 743 '~Spare MB1[23].7'; 744 '~Spare MB1[23].8'; 745 '~Spare MB1[23].9'; 746 '~Spare MB1[23].10'; 747 '~Spare MB1[23].11'; 748 '~Spare MB1[23].12'; 749 '~Spare MB1[23].13'; 750 '~Spare MB1[23].14'; 751 '~Spare MB1[23].15'; 752 '~Spare MB1[23].16'; 753 '~Spare MB1[23].17'; 754 '~Spare MB1[23].18'; 755 '~Spare MB1[23].19'; 756 '~Spare MB1[23].20'; 757 '~Spare MB1[23].21'; 758 '~Spare MB1[23].22'; 759 '~Spare MB1[23].23'; 760 '~Spare MB1[23].24'; 761 '~Spare MB1[23].25'; 762 '~Spare MB1[23].26'; 763 '~Spare MB1[23].27'; 764 '~Spare MB1[23].28'; 765 '~Spare MB1[23].29'; 766 '~Spare MB1[23].30'; 767 '~Spare MB1[23].31'; 768 '~S001R04ES1 - S001R04 EtherNet Switch Connection Inhibited MB1[24].0'; 769 '~Spare MB1[24].1'; 770 '~Spare MB1[24].2'; 771 '~Spare MB1[24].3'; 772 '~Spare MB1[24].4'; 773 '~Spare MB1[24].5'; 774 '~Spare MB1[24].6'; 775 '~Spare MB1[24].7'; 776 '~Spare MB1[24].8'; 777 '~Spare MB1[24].9'; 778 '~Spare MB1[24].10'; 779 '~Spare MB1[24].11'; 780 '~Spare MB1[24].12'; 781 '~Spare MB1[24].13'; 782 '~Spare MB1[24].14'; 783 '~Spare MB1[24].15'; 784 '~Spare MB1[24].16'; 785 '~S001R04Sfty - Robot E-Stop Depressed MB1[24].17'; 786 '~S001R04Sfty - Robot Safety Interface Not Enabled MB1[24].18'; 787 '~S001R04Sfty - Robot DCS Has Been Edited MB1[24].19'; 788 '~S001R04CN - Robot Controller Connection Inhibited MB1[24].20'; 789 '~S001R04E#B# - Robot End Effector Module Connection Inhibited MB1[24].21'; 790 '~S001R04E#B# - Robot End Effector Module Connection Inhibited MB1[24].22'; 791 '~S001R04E#B# - Robot End Effector Module Connection Inhibited MB1[24].23'; 792 '~S001R04E#B# - Robot End Effector Module Connection Inhibited MB1[24].24'; 793 '~S001R04E#B# - Robot End Effector Module Connection Inhibited MB1[24].25'; 794 '~S001R04E#B# - Robot End Effector Module Connection Inhibited MB1[24].26'; 795 '~S001R04E#B# - Robot End Effector Module Connection Inhibited MB1[24].27'; 796 '~S001R04E#B# - Robot End Effector Module Connection Inhibited MB1[24].28'; 797 '~S001R04E#B# - Robot End Effector Module Connection Inhibited MB1[24].29'; 798 '~Spare MB1[24].30'; 799 '~Spare MB1[24].31'; 800 '~Spare MB1[25].0'; 801 '~S001R04F#B# - Robot Process I/O Connection Inhibited MB1[25].1'; 802 '~S001R04F#B# - Robot Process I/O Connection Inhibited MB1[25].2'; 803 '~S001R04F#B# - Robot Process I/O Connection Inhibited MB1[25].3'; 804 '~S001R04F#B# - Robot Process I/O Connection Inhibited MB1[25].4'; 805 '~Spare MB1[25].5'; 806 '~Spare MB1[25].6'; 807 '~Spare MB1[25].7'; 808 '~Spare MB1[25].8'; 809 '~Spare MB1[25].9'; 810 '~S001R04CN.I.Safety - Chain Fault MB1[25].10'; 811 '~S001R04CN.I.AirOn - Robot Air Not On MB1[25].11'; 812 '~S001R04CN.I.RbtAuto - Robot Not in Auto MB1[25].12'; 813 '~S001R04CN.M.InTeach - Robot In Teach MB1[25].13'; 814 '~S001R04CN.I.AtMaintPos - Robot At Maintenace MB1[25].14'; 815 '~S001R04CN.I.RunEnblInterruptAck - Robot In Hold MB1[25].15'; 816 '~S001R04CN.M.MaintPosSeld - Robot Maintenance Selected MB1[25].16'; 817 '~Spare MB1[25].17'; 818 '~Spare MB1[25].18'; 819 '~Spare MB1[25].19'; 820 '~S001R04CN.I.ExtAppCommFlt - Robot Application Communication Fault MB1[25].20'; 821 '~S001R04CN.M.AbortPickupSeld - Robot Abort Pickup Selected MB1[25].21'; 822 '~S001R04CN.M.RetFmPounceSeld - Robot Return From Pounce Selected MB1[25].22'; 823 '~S001R04CN.I.StudWld1 Comm Not OK MB1[25].23'; 824 '~S001R04CN.I.StudWld2 Comm Not OK MB1[25].24'; 825 '~S001R04CN.I.WldMode - Robot In No Weld MB1[25].25'; 826 '~S001R04CN.I.PulledTipBypSS - Robot Pulled Tip Bypass Selected MB1[25].26'; 827 '~S001R04CN.I.FlowNoFlowSS - Robot In No Flow MB1[25].27'; 828 '~S001R04CN.I.RvtNoRvtSS - Robot In No Rivet MB1[25].28'; 829 '~S001R04CN.I.WldCtrlCommOk1 - Robot Weld Controller 1 Comm Not OK MB1[25].29'; 830 '~S001R04CN.I.WldModeStud - Robot In No Weld Stud MB1[25].30'; 831 '~S001R04CN.Ix.MigWldNoWld - Robot In No Weld Mig MB1[25].31'; 832 '~S001R04CN.I.StudWld1Rdy - Robot Stud Weld Controller 1 Not Ready MB1[26].0'; 833 '~S001R04CN.I.Rvt1RdyToOperate - Robot Rivet Controller 1 Not Ready MB1[26].1'; 834 '~S001R04CN.Ix.MigRdy - Robot Mig Weld Controller Not Ready MB1[26].2'; 835 '~S001R04CN.Ix.MigWldNoWld - Robot In No Weld MB1[26].3'; 836 '~Spare MB1[26].4'; 837 '~S001R04CN.I.WldCtrlCommOk2 - Robot Weld Controller 2 Comm Not OK MB1[26].5'; 838 '~Spare MB1[26].6'; 839 '~Spare MB1[26].7'; 840 '~S001R04CN.I.StudWld2Rdy - Robot Stud Weld Controller 2 Not Ready MB1[26].8'; 841 '~S001R04CN.I.Rvt2RdyToOperate - Robot Rivet Controller 2 Not Ready MB1[26].9'; 842 '~S001R04CN.Ix.LaserWldOn - Robot Laser In No Cut MB1[26].10'; 843 '~S001R04CN.Ix.GlassNotPres - Robot Laser Glass Not Present MB1[26].11'; 844 '~S001R04CN.Ix.LaserHeadRdy - Robot Laser Head Not Ready MB1[26].12'; 845 '~S001R04CN.Ix.ChillerOn - Robot Laser Chiller Not On MB1[26].13'; 846 '~S001R04CN.Ix.GasOn - Robot Gas Not On MB1[26].14'; 847 '~S001R04 Power Meter Not Ready MB1[26].15'; 848 '~S001R04 No Wire Present Replace Barrel MB1[26].16'; 849 '~S001R04 Wire Feeder Fault Timer MB1[26].17'; 850 '~S001R04CN.Ix.NRFlt - Robot Nut Runner Not Ready MB1[26].18'; 851 '~Spare MB1[26].19'; 852 '~S001R04CN.M.WrongRivetAtNose - Remove Wrong Rivet At Nose MB1[26].20'; 853 '~S001R04CN.M.DisableRbtDrvs - In Rivet Zone But Riveter Not In Auto MB1[26].21'; 854 '~S001R04CN.I.Rvt1SystemInAuto - Rivet Controller 1 Not In Auto MB1[26].22'; 855 '~S001R04CN.I.Rvt2SystemInAuto - Rivet Controller 2 Not In Auto MB1[26].23'; 856 '~S001R04CN.M.RvtC1ReelCtr.DN - Reel Change Required MB1[26].24'; 857 '~S001R04CN.M.RvtC2ReelCtr.DN - Reel Change Required MB1[26].25'; 858 '~S001R04CN.M.AbortSkipRemain - SkipRemaining Aborted, Reset At Rbt Controller Is Required MB1[26].26'; 859 '~Spare MB1[26].27'; 860 '~Spare MB1[26].28'; 861 '~Spare MB1[26].29'; 862 '~Spare MB1[26].30'; 863 '~Spare MB1[26].31'; 864 '~Spare MB1[27].0'; 865 '~Spare MB1[27].1'; 866 '~Spare MB1[27].2'; 867 '~Spare MB1[27].3'; 868 '~Spare MB1[27].4'; 869 '~Spare MB1[27].5'; 870 '~Spare MB1[27].6'; 871 '~Spare MB1[27].7'; 872 '~Spare MB1[27].8'; 873 '~Spare MB1[27].9'; 874 '~Spare MB1[27].10'; 875 '~Spare MB1[27].11'; 876 '~Spare MB1[27].12'; 877 '~Spare MB1[27].13'; 878 '~Spare MB1[27].14'; 879 '~Spare MB1[27].15'; 880 '~Spare MB1[27].16'; 881 '~Spare MB1[27].17'; 882 '~Spare MB1[27].18'; 883 '~Spare MB1[27].19'; 884 '~Spare MB1[27].20'; 885 '~Spare MB1[27].21'; 886 '~Spare MB1[27].22'; 887 '~Spare MB1[27].23'; 888 '~Spare MB1[27].24'; 889 '~Spare MB1[27].25'; 890 '~Spare MB1[27].26'; 891 '~Spare MB1[27].27'; 892 '~Spare MB1[27].28'; 893 '~Spare MB1[27].29'; 894 '~Spare MB1[27].30'; 895 '~Spare MB1[27].31'; 896 '~Spare MB1[28].0'; 897 '~Spare MB1[28].1'; 898 '~Spare MB1[28].2'; 899 '~Spare MB1[28].3'; 900 '~Spare MB1[28].4'; 901 '~Spare MB1[28].5'; 902 '~Spare MB1[28].6'; 903 '~Spare MB1[28].7'; 904 '~Spare MB1[28].8'; 905 '~Spare MB1[28].9'; 906 '~Spare MB1[28].10'; 907 '~Spare MB1[28].11'; 908 '~Spare MB1[28].12'; 909 '~Spare MB1[28].13'; 910 '~Spare MB1[28].14'; 911 '~Spare MB1[28].15'; 912 '~Spare MB1[28].16'; 913 '~Spare MB1[28].17'; 914 '~Spare MB1[28].18'; 915 '~Spare MB1[28].19'; 916 '~Spare MB1[28].20'; 917 '~Spare MB1[28].21'; 918 '~Spare MB1[28].22'; 919 '~Spare MB1[28].23'; 920 '~Spare MB1[28].24'; 921 '~Spare MB1[28].25'; 922 '~Spare MB1[28].26'; 923 '~Spare MB1[28].27'; 924 '~Spare MB1[28].28'; 925 '~Spare MB1[28].29'; 926 '~Spare MB1[28].30'; 927 '~Spare MB1[28].31'; 928 '~Spare MB1[29].0'; 929 '~Spare MB1[29].1'; 930 '~Spare MB1[29].2'; 931 '~Spare MB1[29].3'; 932 '~Spare MB1[29].4'; 933 '~Spare MB1[29].5'; 934 '~Spare MB1[29].6'; 935 '~Spare MB1[29].7'; 936 '~Spare MB1[29].8'; 937 '~Spare MB1[29].9'; 938 '~Spare MB1[29].10'; 939 '~Spare MB1[29].11'; 940 '~Spare MB1[29].12'; 941 '~Spare MB1[29].13'; 942 '~Spare MB1[29].14'; 943 '~Spare MB1[29].15'; 944 '~Spare MB1[29].16'; 945 '~Spare MB1[29].17'; 946 '~Spare MB1[29].18'; 947 '~Spare MB1[29].19'; 948 '~Spare MB1[29].20'; 949 '~Spare MB1[29].21'; 950 '~Spare MB1[29].22'; 951 '~Spare MB1[29].23'; 952 '~Spare MB1[29].24'; 953 '~Spare MB1[29].25'; 954 '~Spare MB1[29].26'; 955 '~Spare MB1[29].27'; 956 '~Spare MB1[29].28'; 957 '~Spare MB1[29].29'; 958 '~Spare MB1[29].30'; 959 '~Spare MB1[29].31'; 960 '~S001R05ES1 - S001R05 EtherNet Switch Connection Inhibited MB1[30].0'; 961 '~Spare MB1[30].1'; 962 '~Spare MB1[30].2'; 963 '~Spare MB1[30].3'; 964 '~Spare MB1[30].4'; 965 '~Spare MB1[30].5'; 966 '~Spare MB1[30].6'; 967 '~Spare MB1[30].7'; 968 '~Spare MB1[30].8'; 969 '~Spare MB1[30].9'; 970 '~Spare MB1[30].10'; 971 '~Spare MB1[30].11'; 972 '~Spare MB1[30].12'; 973 '~Spare MB1[30].13'; 974 '~Spare MB1[30].14'; 975 '~Spare MB1[30].15'; 976 '~Spare MB1[30].16'; 977 '~S001R05Sfty - Robot E-Stop Depressed MB1[30].17'; 978 '~S001R05Sfty - Robot Safety Interface Not Enabled MB1[30].18'; 979 '~S001R05Sfty - Robot DCS Has Been Edited MB1[30].19'; 980 '~S001R05CN - Robot Controller Connection Inhibited MB1[30].20'; 981 '~S001R05E#B# - Robot End Effector Module Connection Inhibited MB1[30].21'; 982 '~S001R05E#B# - Robot End Effector Module Connection Inhibited MB1[30].22'; 983 '~S001R05E#B# - Robot End Effector Module Connection Inhibited MB1[30].23'; 984 '~S001R05E#B# - Robot End Effector Module Connection Inhibited MB1[30].24'; 985 '~S001R05E#B# - Robot End Effector Module Connection Inhibited MB1[30].25'; 986 '~S001R05E#B# - Robot End Effector Module Connection Inhibited MB1[30].26'; 987 '~S001R05E#B# - Robot End Effector Module Connection Inhibited MB1[30].27'; 988 '~S001R05E#B# - Robot End Effector Module Connection Inhibited MB1[30].28'; 989 '~S001R05E#B# - Robot End Effector Module Connection Inhibited MB1[30].29'; 990 '~Spare MB1[30].30'; 991 '~Spare MB1[30].31'; 992 '~Spare MB1[31].0'; 993 '~S001R05F#B# - Robot Process I/O Connection Inhibited MB1[31].1'; 994 '~S001R05F#B# - Robot Process I/O Connection Inhibited MB1[31].2'; 995 '~S001R05F#B# - Robot Process I/O Connection Inhibited MB1[31].3'; 996 '~S001R05F#B# - Robot Process I/O Connection Inhibited MB1[31].4'; 997 '~Spare MB1[31].5'; 998 '~Spare MB1[31].6'; 999 '~Spare MB1[31].7'; 1000 '~Spare MB1[31].8'; 1001 '~Spare MB1[31].9'; 1002 '~S001R05CN.I.Safety - Chain Fault MB1[31].10'; 1003 '~S001R05CN.I.AirOn - Robot Air Not On MB1[31].11'; 1004 '~S001R05CN.I.RbtAuto - Robot Not in Auto MB1[31].12'; 1005 '~S001R05CN.M.InTeach - Robot In Teach MB1[31].13'; 1006 '~S001R05CN.I.AtMaintPos - Robot At Maintenace MB1[31].14'; 1007 '~S001R05CN.I.RunEnblInterruptAck - Robot In Hold MB1[31].15'; 1008 '~S001R05CN.M.MaintPosSeld - Robot Maintenance Selected MB1[31].16'; 1009 '~Spare MB1[31].17'; 1010 '~Spare MB1[31].18'; 1011 '~Spare MB1[31].19'; 1012 '~S001R05CN.I.ExtAppCommFlt - Robot Application Communication Fault MB1[31].20'; 1013 '~S001R05CN.M.AbortPickupSeld - Robot Abort Pickup Selected MB1[31].21'; 1014 '~S001R05CN.M.RetFmPounceSeld - Robot Return From Pounce Selected MB1[31].22'; 1015 '~S001R05CN.I.StudWld1 Comm Not OK MB1[31].23'; 1016 '~S001R05CN.I.StudWld2 Comm Not OK MB1[31].24'; 1017 '~S001R05CN.I.WldMode - Robot In No Weld MB1[31].25'; 1018 '~S001R05CN.I.PulledTipBypSS - Robot Pulled Tip Bypass Selected MB1[31].26'; 1019 '~S001R05CN.I.FlowNoFlowSS - Robot In No Flow MB1[31].27'; 1020 '~S001R05CN.I.RvtNoRvtSS - Robot In No Rivet MB1[31].28'; 1021 '~S001R05CN.I.WldCtrlCommOk1 - Robot Weld Controller 1 Comm Not OK MB1[31].29'; 1022 '~S001R05CN.I.WldModeStud - Robot In No Weld Stud MB1[31].30'; 1023 '~S001R05CN.Ix.MigWldNoWld - Robot In No Weld Mig MB1[31].31'; 1024 '~S001R05CN.I.StudWld1Rdy - Robot Stud Weld Controller 1 Not Ready MB1[32].0'; 1025 '~S001R05CN.I.Rvt1RdyToOperate - Robot Rivet Controller 1 Not Ready MB1[32].1'; 1026 '~S001R05CN.Ix.MigRdy - Robot Mig Weld Controller Not Ready MB1[32].2'; 1027 